(* Logix 5000 project; controller FV vendor 1 type 14 code 217 rev 31.11; software revision 31.00; part 36 of 63 *)
(* tags used below, declared in another part *)
   Alarm_Reset : BOOL;
   Analog_Fault_No : DINT;
   Analog_Simulation_Enabled : BOOL;
   CWD : CHECKWORD_FLAGS;
   Default_Check_Time : DINT;
   FV_FV10_TTX01_AI : PlantItem;   // FV10_TTX01
   FV_FV10_TTX01_AI_RawInput : ALIAS FOR Remote_IO:11:I.Ch1Data;   // Real Analog Input , Do Not Use In Code
   FV_FV11_TTX01_AI : PlantItem;   // FV11_TTX01
   FV_FV11_TTX01_AI_RawInput : ALIAS FOR Remote_IO:11:I.Ch2Data;   // Real Analog Input , Do Not Use In Code
   FV_FV12_TTX01_AI : PlantItem;   // FV12_TTX01
   FV_FV12_TTX01_AI_RawInput : ALIAS FOR Remote_IO:11:I.Ch3Data;   // Real Analog Input , Do Not Use In Code
   FV_FV13_TTX01_AI : PlantItem;   // FV13_TTX01
   FV_FV13_TTX01_AI_RawInput : ALIAS FOR Remote_IO:11:I.Ch4Data;   // Real Analog Input , Do Not Use In Code
   FV_FV14_TTX01_AI : PlantItem;   // FV14_TTX01
   FV_FV14_TTX01_AI_RawInput : ALIAS FOR Remote_IO:11:I.Ch5Data;   // Real Analog Input , Do Not Use In Code
   FV_FV15_TTX01_AI : PlantItem;   // FV15_TTX01
   FV_FV15_TTX01_AI_RawInput : ALIAS FOR Remote_IO:11:I.Ch6Data;   // Real Analog Input , Do Not Use In Code
   FV_FV16_TTX01_AI : PlantItem;   // FV16_TTX01
   FV_FV16_TTX01_AI_RawInput : ALIAS FOR Remote_IO:11:I.Ch7Data;   // Real Analog Input , Do Not Use In Code
   FV_FV17_TTX01_AI : PlantItem;   // FV17_TTX01
   FV_FV17_TTX01_AI_RawInput : ALIAS FOR Remote_IO:12:I.Ch0Data;   // Real Analog Input , Do Not Use In Code
   FV_FV18_TTX01_AI : PlantItem;   // FV18_TTX01
   FV_FV18_TTX01_AI_RawInput : ALIAS FOR Remote_IO:12:I.Ch1Data;   // Real Analog Input , Do Not Use In Code
   FV_FV19_TTX01_AI : PlantItem;   // FV19_TTX01
   FV_FV19_TTX01_AI_RawInput : ALIAS FOR Remote_IO:12:I.Ch2Data;   // Real Analog Input , Do Not Use In Code
   FV_FV20_TTX01_AI : PlantItem;   // FV20_TTX01
   FV_FV20_TTX01_AI_RawInput : ALIAS FOR Remote_IO:12:I.Ch3Data;   // Real Analog Input , Do Not Use In Code
   FV_FV21_TTX01_AI : PlantItem;   // FV21_TTX01
   FV_FV21_TTX01_AI_RawInput : ALIAS FOR Remote_IO:12:I.Ch4Data;   // Real Analog Input , Do Not Use In Code
   FV_FV22_TTX01_AI : PlantItem;   // FV22_TTX01
   FV_FV22_TTX01_AI_RawInput : ALIAS FOR Remote_IO:12:I.Ch5Data;   // Real Analog Input , Do Not Use In Code
   FV_FV23_TTX01_AI : PlantItem;   // FV23_TTX01
   FV_FV23_TTX01_AI_RawInput : ALIAS FOR Remote_IO:12:I.Ch6Data;   // Real Analog Input , Do Not Use In Code
   FV_FV24_TTX01_AI : PlantItem;   // FV24_TTX01
   FV_FV24_TTX01_AI_RawInput : ALIAS FOR Remote_IO:12:I.Ch7Data;   // Real Analog Input , Do Not Use In Code
   FV_FV25_TTX01_AI : PlantItem;   // FV25_TTX01
   FV_FV25_TTX01_AI_RawInput : ALIAS FOR Remote_IO:13:I.Ch0Data;   // Real Analog Input , Do Not Use In Code
   FV_FV8_TTX01_AI : PlantItem;   // FV8_TTX01
   FV_FV8_TTX01_AI_RawInput : ALIAS FOR Remote_IO:10:I.Ch7Data;   // Real Analog Input , Do Not Use In Code
   FV_FV9_TTX01_AI : PlantItem;   // FV9_TTX01
   FV_FV9_TTX01_AI_RawInput : ALIAS FOR Remote_IO:11:I.Ch0Data;   // Real Analog Input , Do Not Use In Code
   FV_YSV1_TTX01_AI : PlantItem;   // YSV1_TTX01
   FV_YSV1_TTX01_AI_RawInput : ALIAS FOR Remote_IO:13:I.Ch1Data;   // Real Analog Input , Do Not Use In Code
   FV_YSV1_WTX01_AI : PlantItem;   // YSV1_WTX01
   FV_YSV1_WTX01_AI_RawInput : ALIAS FOR Remote_IO:13:I.Ch6Data;   // Real Analog Input , Do Not Use In Code
   FV_YSV2_TTX01_AI : PlantItem;   // YSV2_TTX01
   FV_YSV2_TTX01_AI_RawInput : ALIAS FOR Remote_IO:13:I.Ch2Data;   // Real Analog Input , Do Not Use In Code
   FV_YSV2_WTX01_AI : PlantItem;   // YSV2_WTX01
   FV_YSV2_WTX01_AI_RawInput : ALIAS FOR Remote_IO:13:I.Ch5Data;   // Real Analog Input , Do Not Use In Code
   FV_YSV3_TTX01_AI : PlantItem;   // YSV3_TTX01
   FV_YSV3_TTX01_AI_RawInput : ALIAS FOR Remote_IO:13:I.Ch3Data;   // Real Analog Input , Do Not Use In Code
   FV_YSV3_WTX01_AI : PlantItem;   // YSV3_WTX01
   FV_YSV3_WTX01_AI_RawInput : ALIAS FOR Remote_IO:13:I.Ch4Data;   // Real Analog Input , Do Not Use In Code
   One_Second_One_Scan : ALIAS FOR One_Second_1_scan;
   overrange_RIO_analog_value : REAL;
   underrange_RIO_analog_value : REAL;
(* FV_Common, continued *)

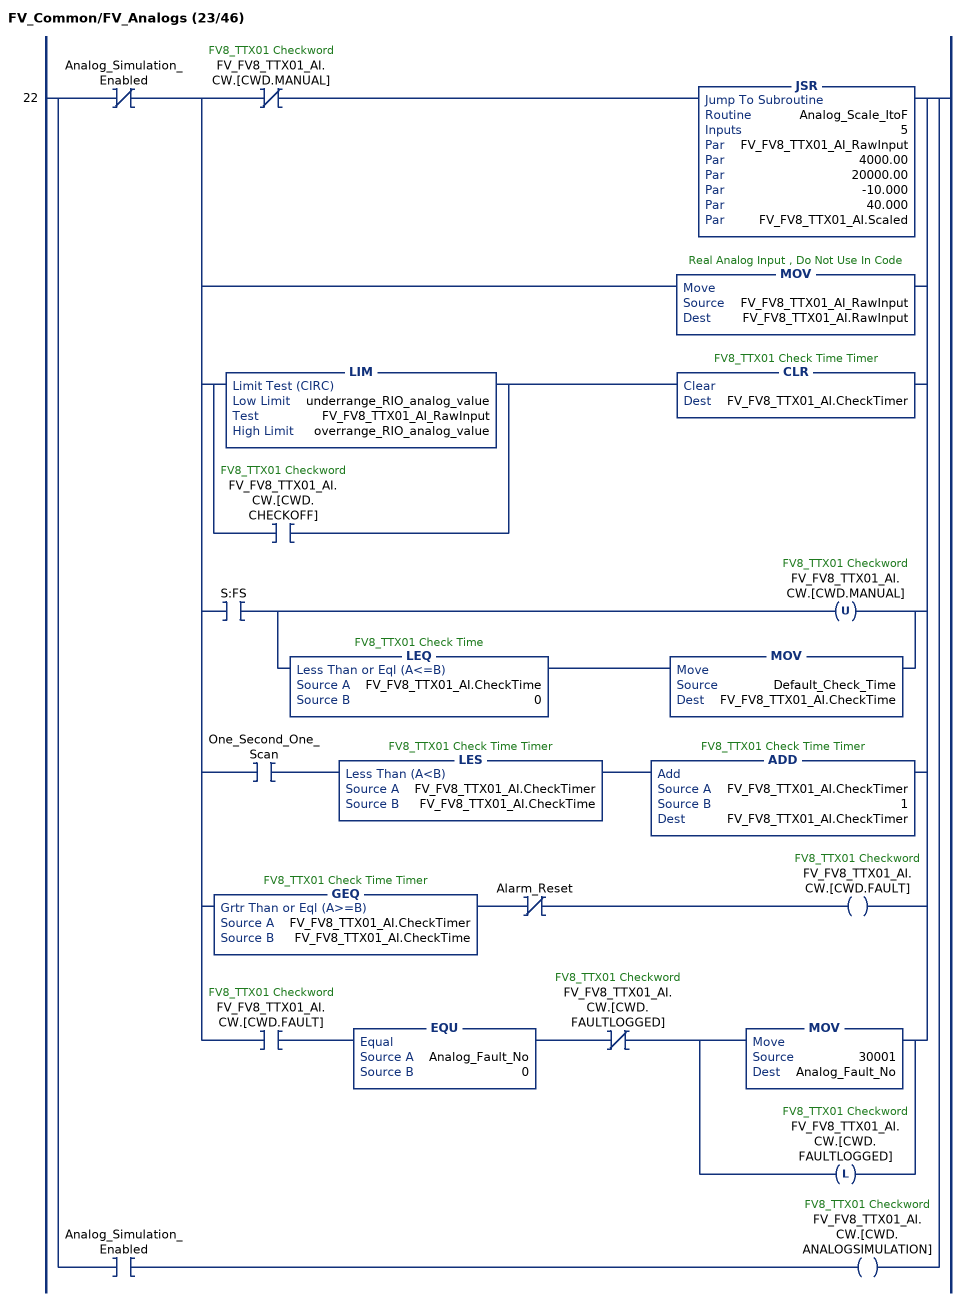
   [picture p757: FV_Common/FV_Analogs rungs 22-22]
   22: [XIO(Analog_Simulation_Enabled) [XIO(FV_FV8_TTX01_AI.CW.[CWD.MANUAL]) JSR(Analog_Scale_ItoF,5,FV_FV8_TTX01_AI_RawInput,4000.00,20000.00,-10.000,40.000,FV_FV8_TTX01_AI.Scaled) ,MOV(FV_FV8_TTX01_AI_RawInput,FV_FV8_TTX01_AI.RawInput) ,[LIM(underrange_RIO_analog_value,FV_FV8_TTX01_AI_RawInput,overrange_RIO_analog_value) ,XIC(FV_FV8_TTX01_AI.CW.[CWD.CHECKOFF]) ] CLR(FV_FV8_TTX01_AI.CheckTimer) ,XIC(S:FS) [OTU(FV_FV8_TTX01_AI.CW.[CWD.MANUAL]) ,LEQ(FV_FV8_TTX01_AI.CheckTime,0) MOV(Default_Check_Time,FV_FV8_TTX01_AI.CheckTime) ] ,XIC(One_Second_One_Scan) LES(FV_FV8_TTX01_AI.CheckTimer,FV_FV8_TTX01_AI.CheckTime) ADD(FV_FV8_TTX01_AI.CheckTimer,1,FV_FV8_TTX01_AI.CheckTimer) ,GEQ(FV_FV8_TTX01_AI.CheckTimer,FV_FV8_TTX01_AI.CheckTime) XIO(Alarm_Reset) OTE(FV_FV8_TTX01_AI.CW.[CWD.FAULT]) ,XIC(FV_FV8_TTX01_AI.CW.[CWD.FAULT]) EQU(Analog_Fault_No,0) XIO(FV_FV8_TTX01_AI.CW.[CWD.FAULTLOGGED]) [MOV(30001,Analog_Fault_No) ,OTL(FV_FV8_TTX01_AI.CW.[CWD.FAULTLOGGED]) ] ] ,XIC(Analog_Simulation_Enabled) OTE(FV_FV8_TTX01_AI.CW.[CWD.ANALOGSIMULATION]) ];
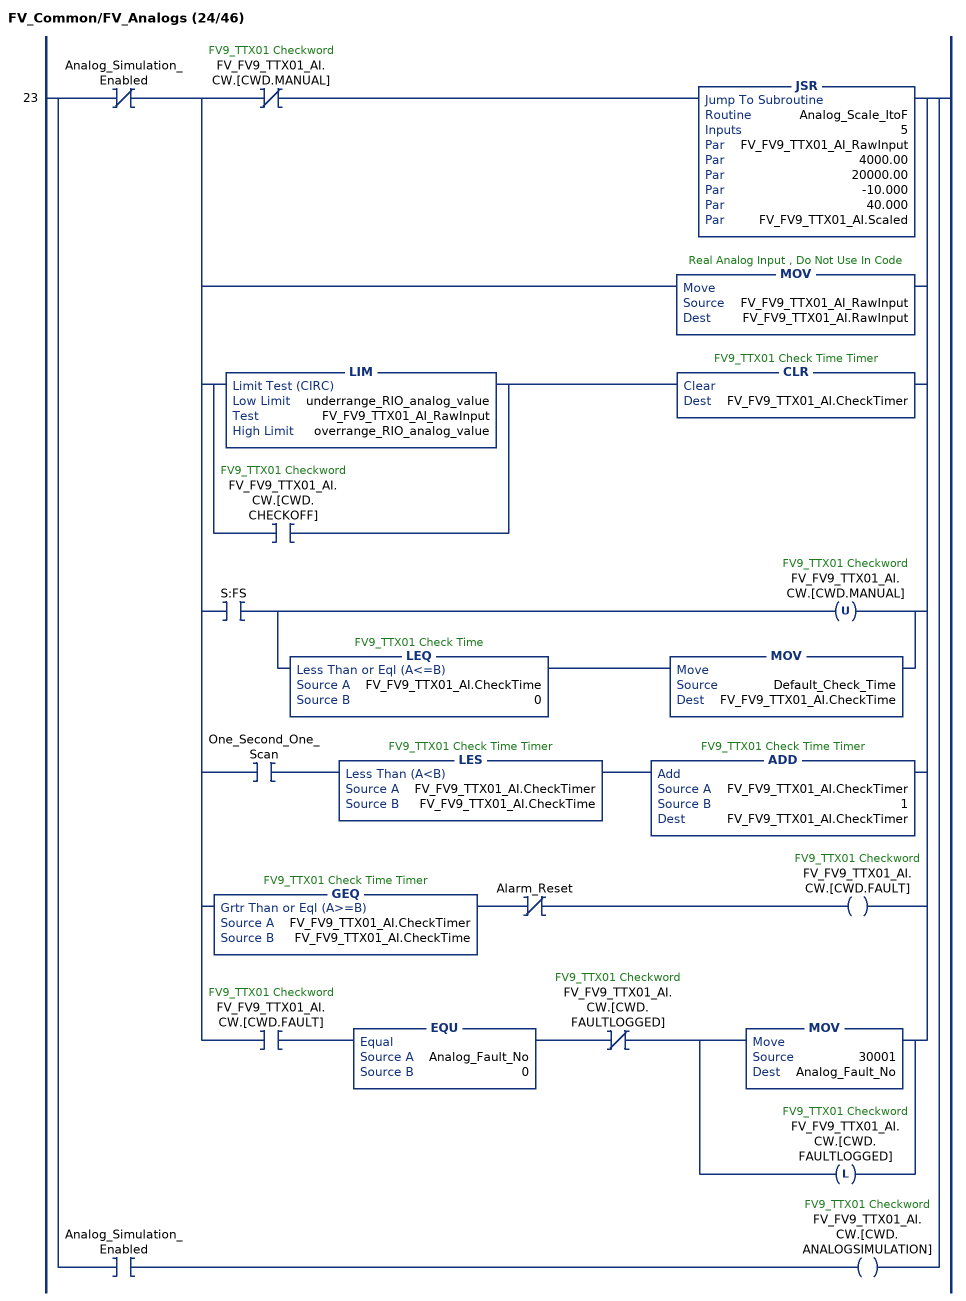
   23: [XIO(Analog_Simulation_Enabled) [XIO(FV_FV9_TTX01_AI.CW.[CWD.MANUAL]) JSR(Analog_Scale_ItoF,5,FV_FV9_TTX01_AI_RawInput,4000.00,20000.00,-10.000,40.000,FV_FV9_TTX01_AI.Scaled) ,MOV(FV_FV9_TTX01_AI_RawInput,FV_FV9_TTX01_AI.RawInput) ,[LIM(underrange_RIO_analog_value,FV_FV9_TTX01_AI_RawInput,overrange_RIO_analog_value) ,XIC(FV_FV9_TTX01_AI.CW.[CWD.CHECKOFF]) ] CLR(FV_FV9_TTX01_AI.CheckTimer) ,XIC(S:FS) [OTU(FV_FV9_TTX01_AI.CW.[CWD.MANUAL]) ,LEQ(FV_FV9_TTX01_AI.CheckTime,0) MOV(Default_Check_Time,FV_FV9_TTX01_AI.CheckTime) ] ,XIC(One_Second_One_Scan) LES(FV_FV9_TTX01_AI.CheckTimer,FV_FV9_TTX01_AI.CheckTime) ADD(FV_FV9_TTX01_AI.CheckTimer,1,FV_FV9_TTX01_AI.CheckTimer) ,GEQ(FV_FV9_TTX01_AI.CheckTimer,FV_FV9_TTX01_AI.CheckTime) XIO(Alarm_Reset) OTE(FV_FV9_TTX01_AI.CW.[CWD.FAULT]) ,XIC(FV_FV9_TTX01_AI.CW.[CWD.FAULT]) EQU(Analog_Fault_No,0) XIO(FV_FV9_TTX01_AI.CW.[CWD.FAULTLOGGED]) [MOV(30001,Analog_Fault_No) ,OTL(FV_FV9_TTX01_AI.CW.[CWD.FAULTLOGGED]) ] ] ,XIC(Analog_Simulation_Enabled) OTE(FV_FV9_TTX01_AI.CW.[CWD.ANALOGSIMULATION]) ];
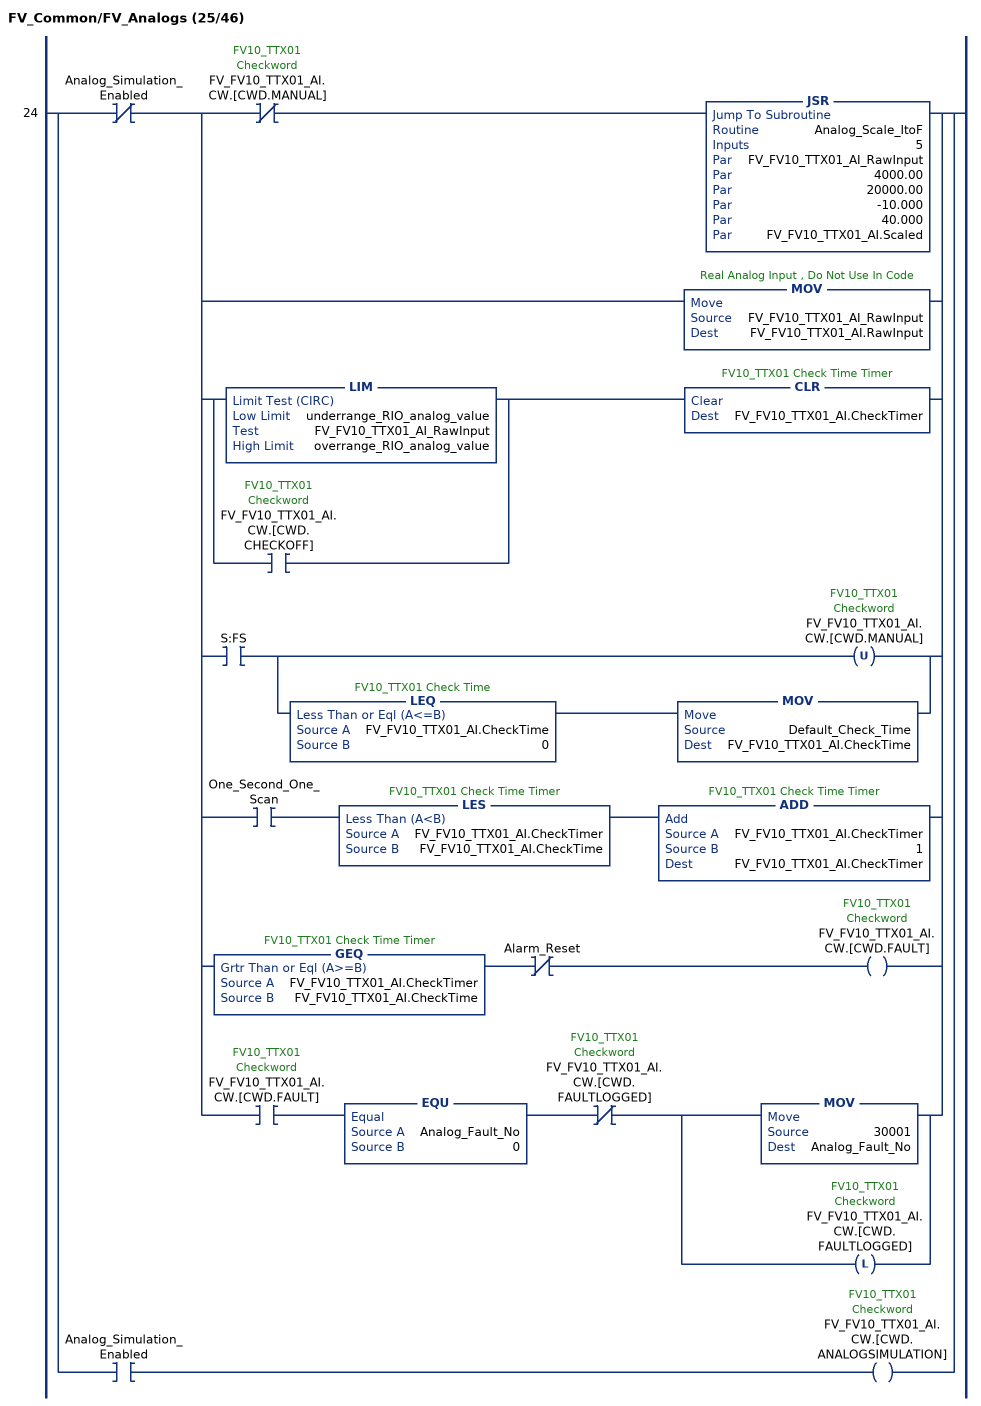
   24: [XIO(Analog_Simulation_Enabled) [XIO(FV_FV10_TTX01_AI.CW.[CWD.MANUAL]) JSR(Analog_Scale_ItoF,5,FV_FV10_TTX01_AI_RawInput,4000.00,20000.00,-10.000,40.000,FV_FV10_TTX01_AI.Scaled) ,MOV(FV_FV10_TTX01_AI_RawInput,FV_FV10_TTX01_AI.RawInput) ,[LIM(underrange_RIO_analog_value,FV_FV10_TTX01_AI_RawInput,overrange_RIO_analog_value) ,XIC(FV_FV10_TTX01_AI.CW.[CWD.CHECKOFF]) ] CLR(FV_FV10_TTX01_AI.CheckTimer) ,XIC(S:FS) [OTU(FV_FV10_TTX01_AI.CW.[CWD.MANUAL]) ,LEQ(FV_FV10_TTX01_AI.CheckTime,0) MOV(Default_Check_Time,FV_FV10_TTX01_AI.CheckTime) ] ,XIC(One_Second_One_Scan) LES(FV_FV10_TTX01_AI.CheckTimer,FV_FV10_TTX01_AI.CheckTime) ADD(FV_FV10_TTX01_AI.CheckTimer,1,FV_FV10_TTX01_AI.CheckTimer) ,GEQ(FV_FV10_TTX01_AI.CheckTimer,FV_FV10_TTX01_AI.CheckTime) XIO(Alarm_Reset) OTE(FV_FV10_TTX01_AI.CW.[CWD.FAULT]) ,XIC(FV_FV10_TTX01_AI.CW.[CWD.FAULT]) EQU(Analog_Fault_No,0) XIO(FV_FV10_TTX01_AI.CW.[CWD.FAULTLOGGED]) [MOV(30001,Analog_Fault_No) ,OTL(FV_FV10_TTX01_AI.CW.[CWD.FAULTLOGGED]) ] ] ,XIC(Analog_Simulation_Enabled) OTE(FV_FV10_TTX01_AI.CW.[CWD.ANALOGSIMULATION]) ];
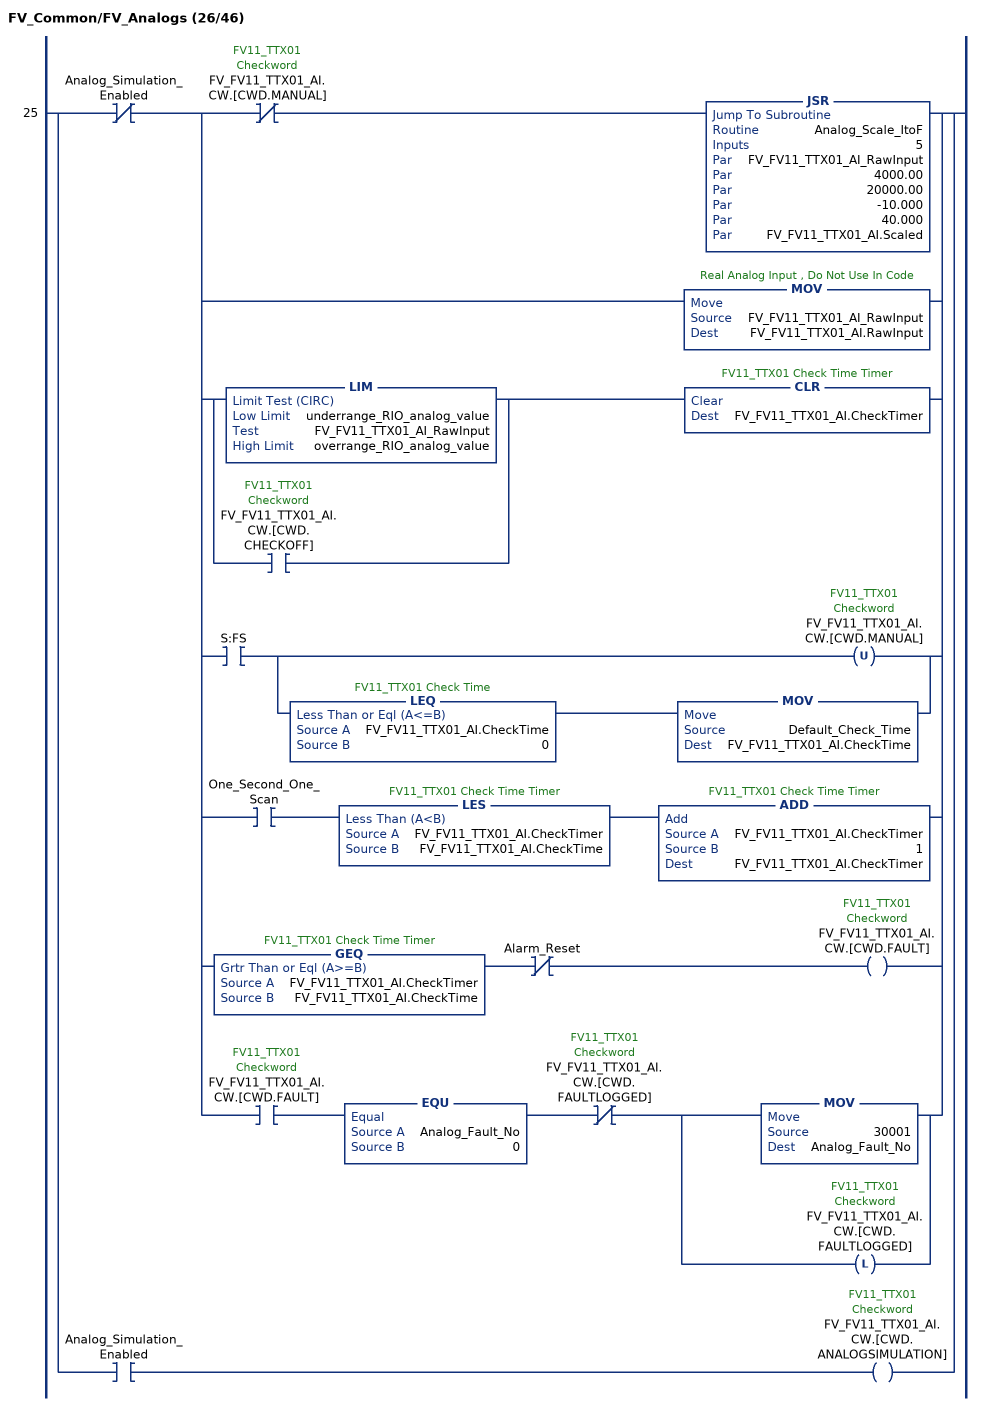
   25: [XIO(Analog_Simulation_Enabled) [XIO(FV_FV11_TTX01_AI.CW.[CWD.MANUAL]) JSR(Analog_Scale_ItoF,5,FV_FV11_TTX01_AI_RawInput,4000.00,20000.00,-10.000,40.000,FV_FV11_TTX01_AI.Scaled) ,MOV(FV_FV11_TTX01_AI_RawInput,FV_FV11_TTX01_AI.RawInput) ,[LIM(underrange_RIO_analog_value,FV_FV11_TTX01_AI_RawInput,overrange_RIO_analog_value) ,XIC(FV_FV11_TTX01_AI.CW.[CWD.CHECKOFF]) ] CLR(FV_FV11_TTX01_AI.CheckTimer) ,XIC(S:FS) [OTU(FV_FV11_TTX01_AI.CW.[CWD.MANUAL]) ,LEQ(FV_FV11_TTX01_AI.CheckTime,0) MOV(Default_Check_Time,FV_FV11_TTX01_AI.CheckTime) ] ,XIC(One_Second_One_Scan) LES(FV_FV11_TTX01_AI.CheckTimer,FV_FV11_TTX01_AI.CheckTime) ADD(FV_FV11_TTX01_AI.CheckTimer,1,FV_FV11_TTX01_AI.CheckTimer) ,GEQ(FV_FV11_TTX01_AI.CheckTimer,FV_FV11_TTX01_AI.CheckTime) XIO(Alarm_Reset) OTE(FV_FV11_TTX01_AI.CW.[CWD.FAULT]) ,XIC(FV_FV11_TTX01_AI.CW.[CWD.FAULT]) EQU(Analog_Fault_No,0) XIO(FV_FV11_TTX01_AI.CW.[CWD.FAULTLOGGED]) [MOV(30001,Analog_Fault_No) ,OTL(FV_FV11_TTX01_AI.CW.[CWD.FAULTLOGGED]) ] ] ,XIC(Analog_Simulation_Enabled) OTE(FV_FV11_TTX01_AI.CW.[CWD.ANALOGSIMULATION]) ];
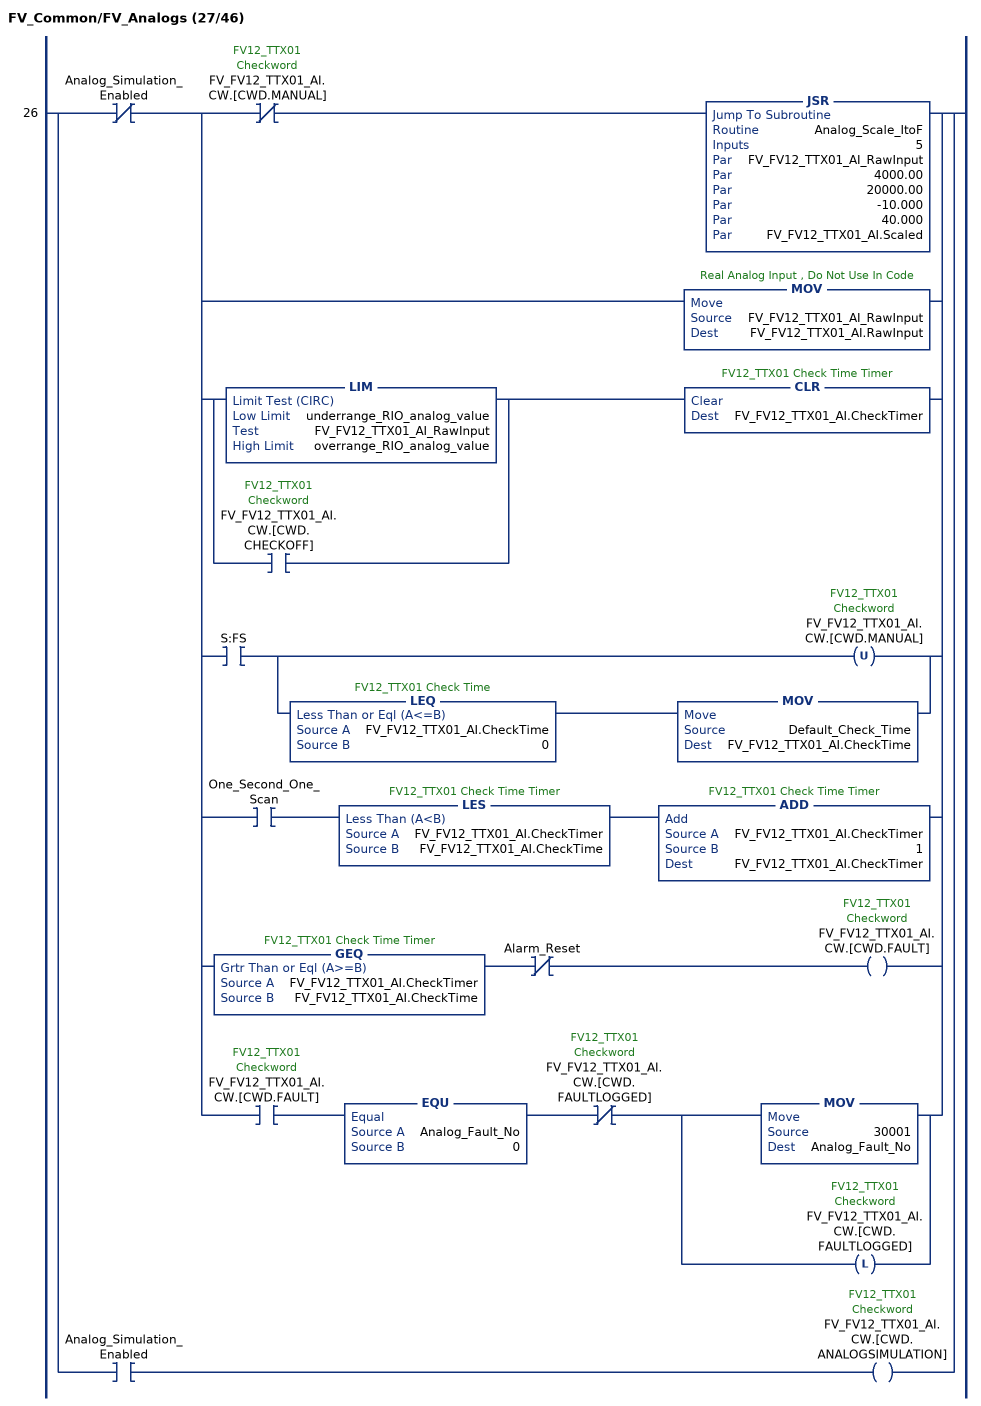
   26: [XIO(Analog_Simulation_Enabled) [XIO(FV_FV12_TTX01_AI.CW.[CWD.MANUAL]) JSR(Analog_Scale_ItoF,5,FV_FV12_TTX01_AI_RawInput,4000.00,20000.00,-10.000,40.000,FV_FV12_TTX01_AI.Scaled) ,MOV(FV_FV12_TTX01_AI_RawInput,FV_FV12_TTX01_AI.RawInput) ,[LIM(underrange_RIO_analog_value,FV_FV12_TTX01_AI_RawInput,overrange_RIO_analog_value) ,XIC(FV_FV12_TTX01_AI.CW.[CWD.CHECKOFF]) ] CLR(FV_FV12_TTX01_AI.CheckTimer) ,XIC(S:FS) [OTU(FV_FV12_TTX01_AI.CW.[CWD.MANUAL]) ,LEQ(FV_FV12_TTX01_AI.CheckTime,0) MOV(Default_Check_Time,FV_FV12_TTX01_AI.CheckTime) ] ,XIC(One_Second_One_Scan) LES(FV_FV12_TTX01_AI.CheckTimer,FV_FV12_TTX01_AI.CheckTime) ADD(FV_FV12_TTX01_AI.CheckTimer,1,FV_FV12_TTX01_AI.CheckTimer) ,GEQ(FV_FV12_TTX01_AI.CheckTimer,FV_FV12_TTX01_AI.CheckTime) XIO(Alarm_Reset) OTE(FV_FV12_TTX01_AI.CW.[CWD.FAULT]) ,XIC(FV_FV12_TTX01_AI.CW.[CWD.FAULT]) EQU(Analog_Fault_No,0) XIO(FV_FV12_TTX01_AI.CW.[CWD.FAULTLOGGED]) [MOV(30001,Analog_Fault_No) ,OTL(FV_FV12_TTX01_AI.CW.[CWD.FAULTLOGGED]) ] ] ,XIC(Analog_Simulation_Enabled) OTE(FV_FV12_TTX01_AI.CW.[CWD.ANALOGSIMULATION]) ];
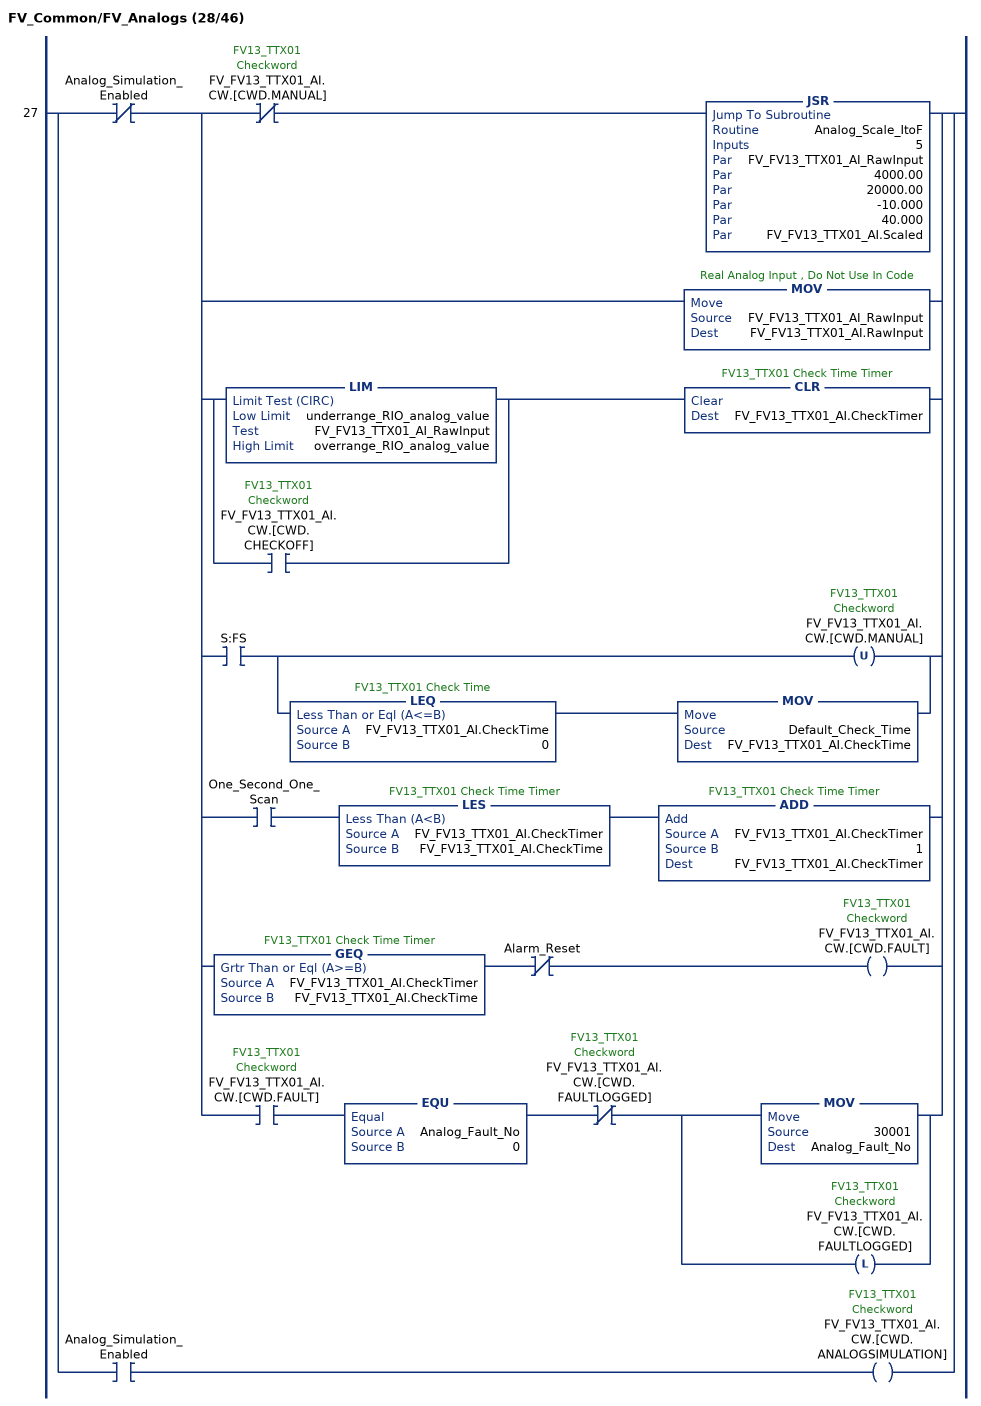
   27: [XIO(Analog_Simulation_Enabled) [XIO(FV_FV13_TTX01_AI.CW.[CWD.MANUAL]) JSR(Analog_Scale_ItoF,5,FV_FV13_TTX01_AI_RawInput,4000.00,20000.00,-10.000,40.000,FV_FV13_TTX01_AI.Scaled) ,MOV(FV_FV13_TTX01_AI_RawInput,FV_FV13_TTX01_AI.RawInput) ,[LIM(underrange_RIO_analog_value,FV_FV13_TTX01_AI_RawInput,overrange_RIO_analog_value) ,XIC(FV_FV13_TTX01_AI.CW.[CWD.CHECKOFF]) ] CLR(FV_FV13_TTX01_AI.CheckTimer) ,XIC(S:FS) [OTU(FV_FV13_TTX01_AI.CW.[CWD.MANUAL]) ,LEQ(FV_FV13_TTX01_AI.CheckTime,0) MOV(Default_Check_Time,FV_FV13_TTX01_AI.CheckTime) ] ,XIC(One_Second_One_Scan) LES(FV_FV13_TTX01_AI.CheckTimer,FV_FV13_TTX01_AI.CheckTime) ADD(FV_FV13_TTX01_AI.CheckTimer,1,FV_FV13_TTX01_AI.CheckTimer) ,GEQ(FV_FV13_TTX01_AI.CheckTimer,FV_FV13_TTX01_AI.CheckTime) XIO(Alarm_Reset) OTE(FV_FV13_TTX01_AI.CW.[CWD.FAULT]) ,XIC(FV_FV13_TTX01_AI.CW.[CWD.FAULT]) EQU(Analog_Fault_No,0) XIO(FV_FV13_TTX01_AI.CW.[CWD.FAULTLOGGED]) [MOV(30001,Analog_Fault_No) ,OTL(FV_FV13_TTX01_AI.CW.[CWD.FAULTLOGGED]) ] ] ,XIC(Analog_Simulation_Enabled) OTE(FV_FV13_TTX01_AI.CW.[CWD.ANALOGSIMULATION]) ];
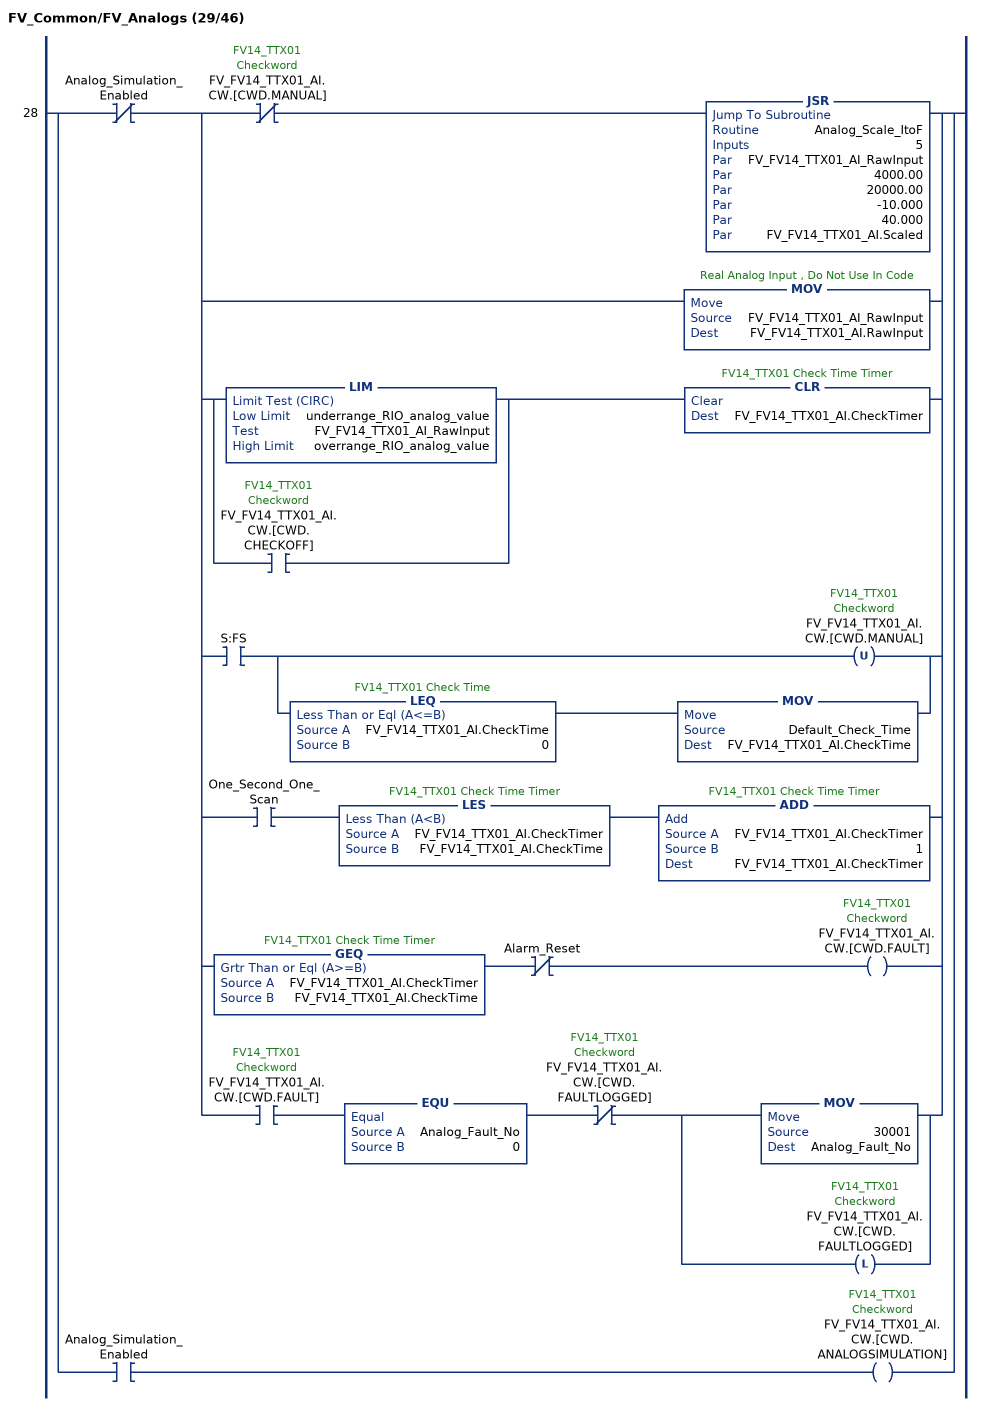
   28: [XIO(Analog_Simulation_Enabled) [XIO(FV_FV14_TTX01_AI.CW.[CWD.MANUAL]) JSR(Analog_Scale_ItoF,5,FV_FV14_TTX01_AI_RawInput,4000.00,20000.00,-10.000,40.000,FV_FV14_TTX01_AI.Scaled) ,MOV(FV_FV14_TTX01_AI_RawInput,FV_FV14_TTX01_AI.RawInput) ,[LIM(underrange_RIO_analog_value,FV_FV14_TTX01_AI_RawInput,overrange_RIO_analog_value) ,XIC(FV_FV14_TTX01_AI.CW.[CWD.CHECKOFF]) ] CLR(FV_FV14_TTX01_AI.CheckTimer) ,XIC(S:FS) [OTU(FV_FV14_TTX01_AI.CW.[CWD.MANUAL]) ,LEQ(FV_FV14_TTX01_AI.CheckTime,0) MOV(Default_Check_Time,FV_FV14_TTX01_AI.CheckTime) ] ,XIC(One_Second_One_Scan) LES(FV_FV14_TTX01_AI.CheckTimer,FV_FV14_TTX01_AI.CheckTime) ADD(FV_FV14_TTX01_AI.CheckTimer,1,FV_FV14_TTX01_AI.CheckTimer) ,GEQ(FV_FV14_TTX01_AI.CheckTimer,FV_FV14_TTX01_AI.CheckTime) XIO(Alarm_Reset) OTE(FV_FV14_TTX01_AI.CW.[CWD.FAULT]) ,XIC(FV_FV14_TTX01_AI.CW.[CWD.FAULT]) EQU(Analog_Fault_No,0) XIO(FV_FV14_TTX01_AI.CW.[CWD.FAULTLOGGED]) [MOV(30001,Analog_Fault_No) ,OTL(FV_FV14_TTX01_AI.CW.[CWD.FAULTLOGGED]) ] ] ,XIC(Analog_Simulation_Enabled) OTE(FV_FV14_TTX01_AI.CW.[CWD.ANALOGSIMULATION]) ];